   3648: 'Spare_Fault_3648', class No Acknowledgement, trigger "DB302_HMI_Faults_Carrier56_Faults_3" bit 15
   3649: 'Carrier 57 Disconnect Open Power Fault DI11.0', class No Acknowledgement, trigger "DB302_HMI_Faults_Carrier57_Faults_0" bit 0
   3650: 'Carrier 57 Drive Profinet Comm Fault', class No Acknowledgement, trigger "DB302_HMI_Faults_Carrier57_Faults_0" bit 1
   3651: 'Carrier 57 Production Stop Not Reset', class No Acknowledgement, trigger "DB302_HMI_Faults_Carrier57_Faults_0" bit 2
   3652: 'Carrier 57 CB02122 Tripped', class No Acknowledgement, trigger "DB302_HMI_Faults_Carrier57_Faults_0" bit 3
   3653: 'Carrier 57 CB02123 Tripped', class No Acknowledgement, trigger "DB302_HMI_Faults_Carrier57_Faults_0" bit 4
   3654: 'Carrier 57 AUX1 CB Tripped', class No Acknowledgement, trigger "DB302_HMI_Faults_Carrier57_Faults_0" bit 5
   3655: 'Carrier 57 AUX2 CB Tripped', class No Acknowledgement, trigger "DB302_HMI_Faults_Carrier57_Faults_0" bit 6
   3656: 'Carrier 57 PLC Not Communicating', class No Acknowledgement, trigger "DB302_HMI_Faults_Carrier57_Faults_0" bit 7
   3657: 'Carrier 57 Safe Input Card Fault', class No Acknowledgement, trigger "DB302_HMI_Faults_Carrier57_Faults_0" bit 8
   3658: 'Carrier 57 Safe Output Card Fault', class No Acknowledgement, trigger "DB302_HMI_Faults_Carrier57_Faults_0" bit 9
   3659: 'Carrier 57 Standard Input Card Fault', class No Acknowledgement, trigger "DB302_HMI_Faults_Carrier57_Faults_0" bit 10
   3660: 'Carrier 57 Standard Output Card Fault', class No Acknowledgement, trigger "DB302_HMI_Faults_Carrier57_Faults_0" bit 11
   3661: 'Carrier 57 Encoder Position Fault', class No Acknowledgement, trigger "DB302_HMI_Faults_Carrier57_Faults_0" bit 12
   3662: 'Carrier 57 Encoder Internal Error', class No Acknowledgement, trigger "DB302_HMI_Faults_Carrier57_Faults_0" bit 13
   3663: 'Carrier 57 Encoder Comm Fault', class No Acknowledgement, trigger "DB302_HMI_Faults_Carrier57_Faults_0" bit 14
   3664: 'Carrier 57 HMI Comm Fault', class No Acknowledgement, trigger "DB302_HMI_Faults_Carrier57_Faults_0" bit 15
   3665: 'Carrier 57 Crash Detection Fault', class No Acknowledgement, trigger "DB302_HMI_Faults_Carrier57_Faults_1" bit 0
   3666: 'Carrier 57 Carrier Number Invalid', class No Acknowledgement, trigger "DB302_HMI_Faults_Carrier57_Faults_1" bit 1
   3667: 'Carrier 57 Drive: PROFINET configuration error', class No Acknowledgement, trigger "DB302_HMI_Faults_Carrier57_Faults_1" bit 2
   3668: 'Carrier 57 Drive: Error internal communications', class No Acknowledgement, trigger "DB302_HMI_Faults_Carrier57_Faults_1" bit 3
   3669: 'Carrier 57 Drive: Motor overtemperature', class No Acknowledgement, trigger "DB302_HMI_Faults_Carrier57_Faults_1" bit 4
   3670: 'Carrier 57 Drive: Motor overcurrent', class No Acknowledgement, trigger "DB302_HMI_Faults_Carrier57_Faults_1" bit 5
   3671: 'Carrier 57 Drive: Infeed or power unit not ready', class No Acknowledgement, trigger "DB302_HMI_Faults_Carrier57_Faults_1" bit 6
   3672: 'Carrier 57 Drive: Short-circuit/ground fault detected', class No Acknowledgement, trigger "DB302_HMI_Faults_Carrier57_Faults_1" bit 7
   3673: 'Carrier 57 Drive: PROFINET Setpoint timeout', class No Acknowledgement, trigger "DB302_HMI_Faults_Carrier57_Faults_1" bit 8
   3674: 'Carrier 57 Power unit: Overcurrent', class No Acknowledgement, trigger "DB302_HMI_Faults_Carrier57_Faults_1" bit 9
   3675: 'Carrier 57 Power unit: DC link voltage overvoltage', class No Acknowledgement, trigger "DB302_HMI_Faults_Carrier57_Faults_1" bit 10
   3676: 'Carrier 57 Power unit: DC link voltage undervoltage', class No Acknowledgement, trigger "DB302_HMI_Faults_Carrier57_Faults_1" bit 11
   3677: 'Carrier 57 Power unit: Line phase failure in main circuit', class No Acknowledgement, trigger "DB302_HMI_Faults_Carrier57_Faults_1" bit 12
   3678: 'Carrier 57 Power unit: Phase failure motor cable', class No Acknowledgement, trigger "DB302_HMI_Faults_Carrier57_Faults_1" bit 13
   3679: 'Carrier 57 Power unit: Ground fault', class No Acknowledgement, trigger "DB302_HMI_Faults_Carrier57_Faults_1" bit 14
   3680: 'Spare_Fault_3680', class No Acknowledgement, trigger "DB302_HMI_Faults_Carrier57_Faults_1" bit 15
   3681: 'Carrier 57 Motion Off Fault', class No Acknowledgement, trigger "DB302_HMI_Faults_Carrier57_Faults_2" bit 0
   3682: 'Carrier 57 Motion On Fault', class No Acknowledgement, trigger "DB302_HMI_Faults_Carrier57_Faults_2" bit 1
   3683: 'Carrier 57 Spacing Fault', class No Acknowledgement, trigger "DB302_HMI_Faults_Carrier57_Faults_2" bit 2
   3684: 'Carrier 57 Duplicate Carrier Number Fault', class No Acknowledgement, trigger "DB302_HMI_Faults_Carrier57_Faults_2" bit 3
   3685: 'Spare_Fault_3685', class No Acknowledgement, trigger "DB302_HMI_Faults_Carrier57_Faults_2" bit 4
   3686: 'Spare_Fault_3686', class No Acknowledgement, trigger "DB302_HMI_Faults_Carrier57_Faults_2" bit 5
   3687: 'Spare_Fault_3687', class No Acknowledgement, trigger "DB302_HMI_Faults_Carrier57_Faults_2" bit 6
   3688: 'Spare_Fault_3688', class No Acknowledgement, trigger "DB302_HMI_Faults_Carrier57_Faults_2" bit 7
   3689: 'Spare_Fault_3689', class No Acknowledgement, trigger "DB302_HMI_Faults_Carrier57_Faults_2" bit 8
   3690: 'Spare_Fault_3690', class No Acknowledgement, trigger "DB302_HMI_Faults_Carrier57_Faults_2" bit 9
   3691: 'Spare_Fault_3691', class No Acknowledgement, trigger "DB302_HMI_Faults_Carrier57_Faults_2" bit 10
   3692: 'Spare_Fault_3692', class No Acknowledgement, trigger "DB302_HMI_Faults_Carrier57_Faults_2" bit 11
   3693: 'Spare_Fault_3693', class No Acknowledgement, trigger "DB302_HMI_Faults_Carrier57_Faults_2" bit 12
   3694: 'Spare_Fault_3694', class No Acknowledgement, trigger "DB302_HMI_Faults_Carrier57_Faults_2" bit 13
   3695: 'Spare_Fault_3695', class No Acknowledgement, trigger "DB302_HMI_Faults_Carrier57_Faults_2" bit 14
   3696: 'Spare_Fault_3696', class No Acknowledgement, trigger "DB302_HMI_Faults_Carrier57_Faults_2" bit 15
   3697: 'Spare_Fault_3697', class No Acknowledgement, trigger "DB302_HMI_Faults_Carrier57_Faults_3" bit 0
   3698: 'Spare_Fault_3698', class No Acknowledgement, trigger "DB302_HMI_Faults_Carrier57_Faults_3" bit 1
   3699: 'Spare_Fault_3699', class No Acknowledgement, trigger "DB302_HMI_Faults_Carrier57_Faults_3" bit 2
   3700: 'Spare_Fault_3700', class No Acknowledgement, trigger "DB302_HMI_Faults_Carrier57_Faults_3" bit 3
   3701: 'Spare_Fault_3701', class No Acknowledgement, trigger "DB302_HMI_Faults_Carrier57_Faults_3" bit 4
   3702: 'Spare_Fault_3702', class No Acknowledgement, trigger "DB302_HMI_Faults_Carrier57_Faults_3" bit 5
   3703: 'Spare_Fault_3703', class No Acknowledgement, trigger "DB302_HMI_Faults_Carrier57_Faults_3" bit 6
   3704: 'Spare_Fault_3704', class No Acknowledgement, trigger "DB302_HMI_Faults_Carrier57_Faults_3" bit 7
   3705: 'Spare_Fault_3705', class No Acknowledgement, trigger "DB302_HMI_Faults_Carrier57_Faults_3" bit 8
   3706: 'Spare_Fault_3706', class No Acknowledgement, trigger "DB302_HMI_Faults_Carrier57_Faults_3" bit 9
   3707: 'Spare_Fault_3707', class No Acknowledgement, trigger "DB302_HMI_Faults_Carrier57_Faults_3" bit 10
   3708: 'Spare_Fault_3708', class No Acknowledgement, trigger "DB302_HMI_Faults_Carrier57_Faults_3" bit 11
   3709: 'Spare_Fault_3709', class No Acknowledgement, trigger "DB302_HMI_Faults_Carrier57_Faults_3" bit 12
   3710: 'Spare_Fault_3710', class No Acknowledgement, trigger "DB302_HMI_Faults_Carrier57_Faults_3" bit 13
   3711: 'Spare_Fault_3711', class No Acknowledgement, trigger "DB302_HMI_Faults_Carrier57_Faults_3" bit 14
   3712: 'Spare_Fault_3712', class No Acknowledgement, trigger "DB302_HMI_Faults_Carrier57_Faults_3" bit 15
   3713: 'Carrier 58 Disconnect Open Power Fault DI11.0', class No Acknowledgement, trigger "DB302_HMI_Faults_Carrier58_Faults_0" bit 0
   3714: 'Carrier 58 Drive Profinet Comm Fault', class No Acknowledgement, trigger "DB302_HMI_Faults_Carrier58_Faults_0" bit 1
   3715: 'Carrier 58 Production Stop Not Reset', class No Acknowledgement, trigger "DB302_HMI_Faults_Carrier58_Faults_0" bit 2
   3716: 'Carrier 58 CB02122 Tripped', class No Acknowledgement, trigger "DB302_HMI_Faults_Carrier58_Faults_0" bit 3
   3717: 'Carrier 58 CB02123 Tripped', class No Acknowledgement, trigger "DB302_HMI_Faults_Carrier58_Faults_0" bit 4
   3718: 'Carrier 58 AUX1 CB Tripped', class No Acknowledgement, trigger "DB302_HMI_Faults_Carrier58_Faults_0" bit 5
   3719: 'Carrier 58 AUX2 CB Tripped', class No Acknowledgement, trigger "DB302_HMI_Faults_Carrier58_Faults_0" bit 6
   3720: 'Carrier 58 PLC Not Communicating', class No Acknowledgement, trigger "DB302_HMI_Faults_Carrier58_Faults_0" bit 7
   3721: 'Carrier 58 Safe Input Card Fault', class No Acknowledgement, trigger "DB302_HMI_Faults_Carrier58_Faults_0" bit 8
   3722: 'Carrier 58 Safe Output Card Fault', class No Acknowledgement, trigger "DB302_HMI_Faults_Carrier58_Faults_0" bit 9
   3723: 'Carrier 58 Standard Input Card Fault', class No Acknowledgement, trigger "DB302_HMI_Faults_Carrier58_Faults_0" bit 10
   3724: 'Carrier 58 Standard Output Card Fault', class No Acknowledgement, trigger "DB302_HMI_Faults_Carrier58_Faults_0" bit 11
   3725: 'Carrier 58 Encoder Position Fault', class No Acknowledgement, trigger "DB302_HMI_Faults_Carrier58_Faults_0" bit 12
   3726: 'Carrier 58 Encoder Internal Error', class No Acknowledgement, trigger "DB302_HMI_Faults_Carrier58_Faults_0" bit 13
   3727: 'Carrier 58 Encoder Comm Fault', class No Acknowledgement, trigger "DB302_HMI_Faults_Carrier58_Faults_0" bit 14
   3728: 'Carrier 58 HMI Comm Fault', class No Acknowledgement, trigger "DB302_HMI_Faults_Carrier58_Faults_0" bit 15
   3729: 'Carrier 58 Crash Detection Fault', class No Acknowledgement, trigger "DB302_HMI_Faults_Carrier58_Faults_1" bit 0
   3730: 'Carrier 58 Carrier Number Invalid', class No Acknowledgement, trigger "DB302_HMI_Faults_Carrier58_Faults_1" bit 1
   3731: 'Carrier 58 Drive: PROFINET configuration error', class No Acknowledgement, trigger "DB302_HMI_Faults_Carrier58_Faults_1" bit 2
   3732: 'Carrier 58 Drive: Error internal communications', class No Acknowledgement, trigger "DB302_HMI_Faults_Carrier58_Faults_1" bit 3
   3733: 'Carrier 58 Drive: Motor overtemperature', class No Acknowledgement, trigger "DB302_HMI_Faults_Carrier58_Faults_1" bit 4
   3734: 'Carrier 58 Drive: Motor overcurrent', class No Acknowledgement, trigger "DB302_HMI_Faults_Carrier58_Faults_1" bit 5
   3735: 'Carrier 58 Drive: Infeed or power unit not ready', class No Acknowledgement, trigger "DB302_HMI_Faults_Carrier58_Faults_1" bit 6
   3736: 'Carrier 58 Drive: Short-circuit/ground fault detected', class No Acknowledgement, trigger "DB302_HMI_Faults_Carrier58_Faults_1" bit 7
   3737: 'Carrier 58 Drive: PROFINET Setpoint timeout', class No Acknowledgement, trigger "DB302_HMI_Faults_Carrier58_Faults_1" bit 8
   3738: 'Carrier 58 Power unit: Overcurrent', class No Acknowledgement, trigger "DB302_HMI_Faults_Carrier58_Faults_1" bit 9
   3739: 'Carrier 58 Power unit: DC link voltage overvoltage', class No Acknowledgement, trigger "DB302_HMI_Faults_Carrier58_Faults_1" bit 10
   3740: 'Carrier 58 Power unit: DC link voltage undervoltage', class No Acknowledgement, trigger "DB302_HMI_Faults_Carrier58_Faults_1" bit 11
   3741: 'Carrier 58 Power unit: Line phase failure in main circuit', class No Acknowledgement, trigger "DB302_HMI_Faults_Carrier58_Faults_1" bit 12
   3742: 'Carrier 58 Power unit: Phase failure motor cable', class No Acknowledgement, trigger "DB302_HMI_Faults_Carrier58_Faults_1" bit 13
   3743: 'Carrier 58 Power unit: Ground fault', class No Acknowledgement, trigger "DB302_HMI_Faults_Carrier58_Faults_1" bit 14
   3744: 'Spare_Fault_3744', class No Acknowledgement, trigger "DB302_HMI_Faults_Carrier58_Faults_1" bit 15
   3745: 'Carrier 58 Motion Off Fault', class No Acknowledgement, trigger "DB302_HMI_Faults_Carrier58_Faults_2" bit 0
   3746: 'Carrier 58 Motion On Fault', class No Acknowledgement, trigger "DB302_HMI_Faults_Carrier58_Faults_2" bit 1
   3747: 'Carrier 58 Spacing Fault', class No Acknowledgement, trigger "DB302_HMI_Faults_Carrier58_Faults_2" bit 2
   3748: 'Carrier 58 Duplicate Carrier Number Fault', class No Acknowledgement, trigger "DB302_HMI_Faults_Carrier58_Faults_2" bit 3
   3749: 'Spare_Fault_3749', class No Acknowledgement, trigger "DB302_HMI_Faults_Carrier58_Faults_2" bit 4
   3750: 'Spare_Fault_3750', class No Acknowledgement, trigger "DB302_HMI_Faults_Carrier58_Faults_2" bit 5
   3751: 'Spare_Fault_3751', class No Acknowledgement, trigger "DB302_HMI_Faults_Carrier58_Faults_2" bit 6
   3752: 'Spare_Fault_3752', class No Acknowledgement, trigger "DB302_HMI_Faults_Carrier58_Faults_2" bit 7
   3753: 'Spare_Fault_3753', class No Acknowledgement, trigger "DB302_HMI_Faults_Carrier58_Faults_2" bit 8
   3754: 'Spare_Fault_3754', class No Acknowledgement, trigger "DB302_HMI_Faults_Carrier58_Faults_2" bit 9
   3755: 'Spare_Fault_3755', class No Acknowledgement, trigger "DB302_HMI_Faults_Carrier58_Faults_2" bit 10
   3756: 'Spare_Fault_3756', class No Acknowledgement, trigger "DB302_HMI_Faults_Carrier58_Faults_2" bit 11
   3757: 'Spare_Fault_3757', class No Acknowledgement, trigger "DB302_HMI_Faults_Carrier58_Faults_2" bit 12
   3758: 'Spare_Fault_3758', class No Acknowledgement, trigger "DB302_HMI_Faults_Carrier58_Faults_2" bit 13
   3759: 'Spare_Fault_3759', class No Acknowledgement, trigger "DB302_HMI_Faults_Carrier58_Faults_2" bit 14
   3760: 'Spare_Fault_3760', class No Acknowledgement, trigger "DB302_HMI_Faults_Carrier58_Faults_2" bit 15
   3761: 'Spare_Fault_3761', class No Acknowledgement, trigger "DB302_HMI_Faults_Carrier58_Faults_3" bit 0
   3762: 'Spare_Fault_3762', class No Acknowledgement, trigger "DB302_HMI_Faults_Carrier58_Faults_3" bit 1
   3763: 'Spare_Fault_3763', class No Acknowledgement, trigger "DB302_HMI_Faults_Carrier58_Faults_3" bit 2
   3764: 'Spare_Fault_3764', class No Acknowledgement, trigger "DB302_HMI_Faults_Carrier58_Faults_3" bit 3
   3765: 'Spare_Fault_3765', class No Acknowledgement, trigger "DB302_HMI_Faults_Carrier58_Faults_3" bit 4
   3766: 'Spare_Fault_3766', class No Acknowledgement, trigger "DB302_HMI_Faults_Carrier58_Faults_3" bit 5
   3767: 'Spare_Fault_3767', class No Acknowledgement, trigger "DB302_HMI_Faults_Carrier58_Faults_3" bit 6
   3768: 'Spare_Fault_3768', class No Acknowledgement, trigger "DB302_HMI_Faults_Carrier58_Faults_3" bit 7
   3769: 'Spare_Fault_3769', class No Acknowledgement, trigger "DB302_HMI_Faults_Carrier58_Faults_3" bit 8
   3770: 'Spare_Fault_3770', class No Acknowledgement, trigger "DB302_HMI_Faults_Carrier58_Faults_3" bit 9
   3771: 'Spare_Fault_3771', class No Acknowledgement, trigger "DB302_HMI_Faults_Carrier58_Faults_3" bit 10
   3772: 'Spare_Fault_3772', class No Acknowledgement, trigger "DB302_HMI_Faults_Carrier58_Faults_3" bit 11
   3773: 'Spare_Fault_3773', class No Acknowledgement, trigger "DB302_HMI_Faults_Carrier58_Faults_3" bit 12
   3774: 'Spare_Fault_3774', class No Acknowledgement, trigger "DB302_HMI_Faults_Carrier58_Faults_3" bit 13
   3775: 'Spare_Fault_3775', class No Acknowledgement, trigger "DB302_HMI_Faults_Carrier58_Faults_3" bit 14
   3776: 'Spare_Fault_3776', class No Acknowledgement, trigger "DB302_HMI_Faults_Carrier58_Faults_3" bit 15
   3777: 'Carrier 59 Disconnect Open Power Fault DI11.0', class No Acknowledgement, trigger "DB302_HMI_Faults_Carrier59_Faults_0" bit 0
   3778: 'Carrier 59 Drive Profinet Comm Fault', class No Acknowledgement, trigger "DB302_HMI_Faults_Carrier59_Faults_0" bit 1
   3779: 'Carrier 59 Production Stop Not Reset', class No Acknowledgement, trigger "DB302_HMI_Faults_Carrier59_Faults_0" bit 2
   3780: 'Carrier 59 CB02122 Tripped', class No Acknowledgement, trigger "DB302_HMI_Faults_Carrier59_Faults_0" bit 3
   3781: 'Carrier 59 CB02123 Tripped', class No Acknowledgement, trigger "DB302_HMI_Faults_Carrier59_Faults_0" bit 4
   3782: 'Carrier 59 AUX1 CB Tripped', class No Acknowledgement, trigger "DB302_HMI_Faults_Carrier59_Faults_0" bit 5
   3783: 'Carrier 59 AUX2 CB Tripped', class No Acknowledgement, trigger "DB302_HMI_Faults_Carrier59_Faults_0" bit 6
   3784: 'Carrier 59 PLC Not Communicating', class No Acknowledgement, trigger "DB302_HMI_Faults_Carrier59_Faults_0" bit 7
   3785: 'Carrier 59 Safe Input Card Fault', class No Acknowledgement, trigger "DB302_HMI_Faults_Carrier59_Faults_0" bit 8
   3786: 'Carrier 59 Safe Output Card Fault', class No Acknowledgement, trigger "DB302_HMI_Faults_Carrier59_Faults_0" bit 9
   3787: 'Carrier 59 Standard Input Card Fault', class No Acknowledgement, trigger "DB302_HMI_Faults_Carrier59_Faults_0" bit 10
   3788: 'Carrier 59 Standard Output Card Fault', class No Acknowledgement, trigger "DB302_HMI_Faults_Carrier59_Faults_0" bit 11
   3789: 'Carrier 59 Encoder Position Fault', class No Acknowledgement, trigger "DB302_HMI_Faults_Carrier59_Faults_0" bit 12
   3790: 'Carrier 59 Encoder Internal Error', class No Acknowledgement, trigger "DB302_HMI_Faults_Carrier59_Faults_0" bit 13
   3791: 'Carrier 59 Encoder Comm Fault', class No Acknowledgement, trigger "DB302_HMI_Faults_Carrier59_Faults_0" bit 14
   3792: 'Carrier 59 HMI Comm Fault', class No Acknowledgement, trigger "DB302_HMI_Faults_Carrier59_Faults_0" bit 15
   3793: 'Carrier 59 Crash Detection Fault', class No Acknowledgement, trigger "DB302_HMI_Faults_Carrier59_Faults_1" bit 0
   3794: 'Carrier 59 Carrier Number Invalid', class No Acknowledgement, trigger "DB302_HMI_Faults_Carrier59_Faults_1" bit 1
   3795: 'Carrier 59 Drive: PROFINET configuration error', class No Acknowledgement, trigger "DB302_HMI_Faults_Carrier59_Faults_1" bit 2
   3796: 'Carrier 59 Drive: Error internal communications', class No Acknowledgement, trigger "DB302_HMI_Faults_Carrier59_Faults_1" bit 3
   3797: 'Carrier 59 Drive: Motor overtemperature', class No Acknowledgement, trigger "DB302_HMI_Faults_Carrier59_Faults_1" bit 4
   3798: 'Carrier 59 Drive: Motor overcurrent', class No Acknowledgement, trigger "DB302_HMI_Faults_Carrier59_Faults_1" bit 5
   3799: 'Carrier 59 Drive: Infeed or power unit not ready', class No Acknowledgement, trigger "DB302_HMI_Faults_Carrier59_Faults_1" bit 6
   3800: 'Carrier 59 Drive: Short-circuit/ground fault detected', class No Acknowledgement, trigger "DB302_HMI_Faults_Carrier59_Faults_1" bit 7
   3801: 'Carrier 59 Drive: PROFINET Setpoint timeout', class No Acknowledgement, trigger "DB302_HMI_Faults_Carrier59_Faults_1" bit 8
   3802: 'Carrier 59 Power unit: Overcurrent', class No Acknowledgement, trigger "DB302_HMI_Faults_Carrier59_Faults_1" bit 9
   3803: 'Carrier 59 Power unit: DC link voltage overvoltage', class No Acknowledgement, trigger "DB302_HMI_Faults_Carrier59_Faults_1" bit 10
   3804: 'Carrier 59 Power unit: DC link voltage undervoltage', class No Acknowledgement, trigger "DB302_HMI_Faults_Carrier59_Faults_1" bit 11
   3805: 'Carrier 59 Power unit: Line phase failure in main circuit', class No Acknowledgement, trigger "DB302_HMI_Faults_Carrier59_Faults_1" bit 12
   3806: 'Carrier 59 Power unit: Phase failure motor cable', class No Acknowledgement, trigger "DB302_HMI_Faults_Carrier59_Faults_1" bit 13
   3807: 'Carrier 59 Power unit: Ground fault', class No Acknowledgement, trigger "DB302_HMI_Faults_Carrier59_Faults_1" bit 14
   3808: 'Spare_Fault_3808', class No Acknowledgement, trigger "DB302_HMI_Faults_Carrier59_Faults_1" bit 15
   3809: 'Carrier 59 Motion Off Fault', class No Acknowledgement, trigger "DB302_HMI_Faults_Carrier59_Faults_2" bit 0
   3810: 'Carrier 59 Motion On Fault', class No Acknowledgement, trigger "DB302_HMI_Faults_Carrier59_Faults_2" bit 1
   3811: 'Carrier 59 Spacing Fault', class No Acknowledgement, trigger "DB302_HMI_Faults_Carrier59_Faults_2" bit 2
   3812: 'Carrier 59 Duplicate Carrier Number Fault', class No Acknowledgement, trigger "DB302_HMI_Faults_Carrier59_Faults_2" bit 3
   3813: 'Spare_Fault_3813', class No Acknowledgement, trigger "DB302_HMI_Faults_Carrier59_Faults_2" bit 4
   3814: 'Spare_Fault_3814', class No Acknowledgement, trigger "DB302_HMI_Faults_Carrier59_Faults_2" bit 5
   3815: 'Spare_Fault_3815', class No Acknowledgement, trigger "DB302_HMI_Faults_Carrier59_Faults_2" bit 6
   3816: 'Spare_Fault_3816', class No Acknowledgement, trigger "DB302_HMI_Faults_Carrier59_Faults_2" bit 7
   3817: 'Spare_Fault_3817', class No Acknowledgement, trigger "DB302_HMI_Faults_Carrier59_Faults_2" bit 8
   3818: 'Spare_Fault_3818', class No Acknowledgement, trigger "DB302_HMI_Faults_Carrier59_Faults_2" bit 9
   3819: 'Spare_Fault_3819', class No Acknowledgement, trigger "DB302_HMI_Faults_Carrier59_Faults_2" bit 10
   3820: 'Spare_Fault_3820', class No Acknowledgement, trigger "DB302_HMI_Faults_Carrier59_Faults_2" bit 11
   3821: 'Spare_Fault_3821', class No Acknowledgement, trigger "DB302_HMI_Faults_Carrier59_Faults_2" bit 12
   3822: 'Spare_Fault_3822', class No Acknowledgement, trigger "DB302_HMI_Faults_Carrier59_Faults_2" bit 13
   3823: 'Spare_Fault_3823', class No Acknowledgement, trigger "DB302_HMI_Faults_Carrier59_Faults_2" bit 14
   3824: 'Spare_Fault_3824', class No Acknowledgement, trigger "DB302_HMI_Faults_Carrier59_Faults_2" bit 15
   3825: 'Spare_Fault_3825', class No Acknowledgement, trigger "DB302_HMI_Faults_Carrier59_Faults_3" bit 0
   3826: 'Spare_Fault_3826', class No Acknowledgement, trigger "DB302_HMI_Faults_Carrier59_Faults_3" bit 1
   3827: 'Spare_Fault_3827', class No Acknowledgement, trigger "DB302_HMI_Faults_Carrier59_Faults_3" bit 2
   3828: 'Spare_Fault_3828', class No Acknowledgement, trigger "DB302_HMI_Faults_Carrier59_Faults_3" bit 3
   3829: 'Spare_Fault_3829', class No Acknowledgement, trigger "DB302_HMI_Faults_Carrier59_Faults_3" bit 4
   3830: 'Spare_Fault_3830', class No Acknowledgement, trigger "DB302_HMI_Faults_Carrier59_Faults_3" bit 5
   3831: 'Spare_Fault_3831', class No Acknowledgement, trigger "DB302_HMI_Faults_Carrier59_Faults_3" bit 6
   3832: 'Spare_Fault_3832', class No Acknowledgement, trigger "DB302_HMI_Faults_Carrier59_Faults_3" bit 7
   3833: 'Spare_Fault_3833', class No Acknowledgement, trigger "DB302_HMI_Faults_Carrier59_Faults_3" bit 8
   3834: 'Spare_Fault_3834', class No Acknowledgement, trigger "DB302_HMI_Faults_Carrier59_Faults_3" bit 9
   3835: 'Spare_Fault_3835', class No Acknowledgement, trigger "DB302_HMI_Faults_Carrier59_Faults_3" bit 10
   3836: 'Spare_Fault_3836', class No Acknowledgement, trigger "DB302_HMI_Faults_Carrier59_Faults_3" bit 11
   3837: 'Spare_Fault_3837', class No Acknowledgement, trigger "DB302_HMI_Faults_Carrier59_Faults_3" bit 12
   3838: 'Spare_Fault_3838', class No Acknowledgement, trigger "DB302_HMI_Faults_Carrier59_Faults_3" bit 13
   3839: 'Spare_Fault_3839', class No Acknowledgement, trigger "DB302_HMI_Faults_Carrier59_Faults_3" bit 14
   3840: 'Spare_Fault_3840', class No Acknowledgement, trigger "DB302_HMI_Faults_Carrier59_Faults_3" bit 15
   3841: 'Carrier 60 Disconnect Open Power Fault DI11.0', class No Acknowledgement, trigger "DB302_HMI_Faults_Carrier60_Faults_0" bit 0
   3842: 'Carrier 60 Drive Profinet Comm Fault', class No Acknowledgement, trigger "DB302_HMI_Faults_Carrier60_Faults_0" bit 1
   3843: 'Carrier 60 Production Stop Not Reset', class No Acknowledgement, trigger "DB302_HMI_Faults_Carrier60_Faults_0" bit 2
   3844: 'Carrier 60 CB02122 Tripped', class No Acknowledgement, trigger "DB302_HMI_Faults_Carrier60_Faults_0" bit 3
   3845: 'Carrier 60 CB02123 Tripped', class No Acknowledgement, trigger "DB302_HMI_Faults_Carrier60_Faults_0" bit 4
   3846: 'Carrier 60 AUX1 CB Tripped', class No Acknowledgement, trigger "DB302_HMI_Faults_Carrier60_Faults_0" bit 5
   3847: 'Carrier 60 AUX2 CB Tripped', class No Acknowledgement, trigger "DB302_HMI_Faults_Carrier60_Faults_0" bit 6
   3848: 'Carrier 60 PLC Not Communicating', class No Acknowledgement, trigger "DB302_HMI_Faults_Carrier60_Faults_0" bit 7
   3849: 'Carrier 60 Safe Input Card Fault', class No Acknowledgement, trigger "DB302_HMI_Faults_Carrier60_Faults_0" bit 8
   3850: 'Carrier 60 Safe Output Card Fault', class No Acknowledgement, trigger "DB302_HMI_Faults_Carrier60_Faults_0" bit 9
   3851: 'Carrier 60 Standard Input Card Fault', class No Acknowledgement, trigger "DB302_HMI_Faults_Carrier60_Faults_0" bit 10
   3852: 'Carrier 60 Standard Output Card Fault', class No Acknowledgement, trigger "DB302_HMI_Faults_Carrier60_Faults_0" bit 11
   3853: 'Carrier 60 Encoder Position Fault', class No Acknowledgement, trigger "DB302_HMI_Faults_Carrier60_Faults_0" bit 12
   3854: 'Carrier 60 Encoder Internal Error', class No Acknowledgement, trigger "DB302_HMI_Faults_Carrier60_Faults_0" bit 13
   3855: 'Carrier 60 Encoder Comm Fault', class No Acknowledgement, trigger "DB302_HMI_Faults_Carrier60_Faults_0" bit 14
   3856: 'Carrier 60 HMI Comm Fault', class No Acknowledgement, trigger "DB302_HMI_Faults_Carrier60_Faults_0" bit 15
   3857: 'Carrier 60 Crash Detection Fault', class No Acknowledgement, trigger "DB302_HMI_Faults_Carrier60_Faults_1" bit 0
   3858: 'Carrier 60 Carrier Number Invalid', class No Acknowledgement, trigger "DB302_HMI_Faults_Carrier60_Faults_1" bit 1
   3859: 'Carrier 60 Drive: PROFINET configuration error', class No Acknowledgement, trigger "DB302_HMI_Faults_Carrier60_Faults_1" bit 2
   3860: 'Carrier 60 Drive: Error internal communications', class No Acknowledgement, trigger "DB302_HMI_Faults_Carrier60_Faults_1" bit 3
   3861: 'Carrier 60 Drive: Motor overtemperature', class No Acknowledgement, trigger "DB302_HMI_Faults_Carrier60_Faults_1" bit 4
   3862: 'Carrier 60 Drive: Motor overcurrent', class No Acknowledgement, trigger "DB302_HMI_Faults_Carrier60_Faults_1" bit 5
   3863: 'Carrier 60 Drive: Infeed or power unit not ready', class No Acknowledgement, trigger "DB302_HMI_Faults_Carrier60_Faults_1" bit 6
   3864: 'Carrier 60 Drive: Short-circuit/ground fault detected', class No Acknowledgement, trigger "DB302_HMI_Faults_Carrier60_Faults_1" bit 7
   3865: 'Carrier 60 Drive: PROFINET Setpoint timeout', class No Acknowledgement, trigger "DB302_HMI_Faults_Carrier60_Faults_1" bit 8
   3866: 'Carrier 60 Power unit: Overcurrent', class No Acknowledgement, trigger "DB302_HMI_Faults_Carrier60_Faults_1" bit 9
   3867: 'Carrier 60 Power unit: DC link voltage overvoltage', class No Acknowledgement, trigger "DB302_HMI_Faults_Carrier60_Faults_1" bit 10
   3868: 'Carrier 60 Power unit: DC link voltage undervoltage', class No Acknowledgement, trigger "DB302_HMI_Faults_Carrier60_Faults_1" bit 11
   3869: 'Carrier 60 Power unit: Line phase failure in main circuit', class No Acknowledgement, trigger "DB302_HMI_Faults_Carrier60_Faults_1" bit 12
   3870: 'Carrier 60 Power unit: Phase failure motor cable', class No Acknowledgement, trigger "DB302_HMI_Faults_Carrier60_Faults_1" bit 13
   3871: 'Carrier 60 Power unit: Ground fault', class No Acknowledgement, trigger "DB302_HMI_Faults_Carrier60_Faults_1" bit 14
   3872: 'Spare_Fault_3872', class No Acknowledgement, trigger "DB302_HMI_Faults_Carrier60_Faults_1" bit 15
   3873: 'Carrier 60 Motion Off Fault', class No Acknowledgement, trigger "DB302_HMI_Faults_Carrier60_Faults_2" bit 0
   3874: 'Carrier 60 Motion On Fault', class No Acknowledgement, trigger "DB302_HMI_Faults_Carrier60_Faults_2" bit 1
   3875: 'Carrier 60 Spacing Fault', class No Acknowledgement, trigger "DB302_HMI_Faults_Carrier60_Faults_2" bit 2
   3876: 'Carrier 60 Duplicate Carrier Number Fault', class No Acknowledgement, trigger "DB302_HMI_Faults_Carrier60_Faults_2" bit 3
   3877: 'Spare_Fault_3877', class No Acknowledgement, trigger "DB302_HMI_Faults_Carrier60_Faults_2" bit 4
   3878: 'Spare_Fault_3878', class No Acknowledgement, trigger "DB302_HMI_Faults_Carrier60_Faults_2" bit 5
   3879: 'Spare_Fault_3879', class No Acknowledgement, trigger "DB302_HMI_Faults_Carrier60_Faults_2" bit 6
   3880: 'Spare_Fault_3880', class No Acknowledgement, trigger "DB302_HMI_Faults_Carrier60_Faults_2" bit 7
   3881: 'Spare_Fault_3881', class No Acknowledgement, trigger "DB302_HMI_Faults_Carrier60_Faults_2" bit 8
   3882: 'Spare_Fault_3882', class No Acknowledgement, trigger "DB302_HMI_Faults_Carrier60_Faults_2" bit 9
   3883: 'Spare_Fault_3883', class No Acknowledgement, trigger "DB302_HMI_Faults_Carrier60_Faults_2" bit 10
   3884: 'Spare_Fault_3884', class No Acknowledgement, trigger "DB302_HMI_Faults_Carrier60_Faults_2" bit 11
   3885: 'Spare_Fault_3885', class No Acknowledgement, trigger "DB302_HMI_Faults_Carrier60_Faults_2" bit 12
   3886: 'Spare_Fault_3886', class No Acknowledgement, trigger "DB302_HMI_Faults_Carrier60_Faults_2" bit 13
   3887: 'Spare_Fault_3887', class No Acknowledgement, trigger "DB302_HMI_Faults_Carrier60_Faults_2" bit 14
   3888: 'Spare_Fault_3888', class No Acknowledgement, trigger "DB302_HMI_Faults_Carrier60_Faults_2" bit 15
   3889: 'Spare_Fault_3889', class No Acknowledgement, trigger "DB302_HMI_Faults_Carrier60_Faults_3" bit 0
   3890: 'Spare_Fault_3890', class No Acknowledgement, trigger "DB302_HMI_Faults_Carrier60_Faults_3" bit 1
   3891: 'Spare_Fault_3891', class No Acknowledgement, trigger "DB302_HMI_Faults_Carrier60_Faults_3" bit 2
   3892: 'Spare_Fault_3892', class No Acknowledgement, trigger "DB302_HMI_Faults_Carrier60_Faults_3" bit 3
   3893: 'Spare_Fault_3893', class No Acknowledgement, trigger "DB302_HMI_Faults_Carrier60_Faults_3" bit 4
   3894: 'Spare_Fault_3894', class No Acknowledgement, trigger "DB302_HMI_Faults_Carrier60_Faults_3" bit 5
   3895: 'Spare_Fault_3895', class No Acknowledgement, trigger "DB302_HMI_Faults_Carrier60_Faults_3" bit 6
   3896: 'Spare_Fault_3896', class No Acknowledgement, trigger "DB302_HMI_Faults_Carrier60_Faults_3" bit 7
   3897: 'Spare_Fault_3897', class No Acknowledgement, trigger "DB302_HMI_Faults_Carrier60_Faults_3" bit 8
   3898: 'Spare_Fault_3898', class No Acknowledgement, trigger "DB302_HMI_Faults_Carrier60_Faults_3" bit 9
   3899: 'Spare_Fault_3899', class No Acknowledgement, trigger "DB302_HMI_Faults_Carrier60_Faults_3" bit 10
   3900: 'Spare_Fault_3900', class No Acknowledgement, trigger "DB302_HMI_Faults_Carrier60_Faults_3" bit 11
   3901: 'Spare_Fault_3901', class No Acknowledgement, trigger "DB302_HMI_Faults_Carrier60_Faults_3" bit 12
   3902: 'Spare_Fault_3902', class No Acknowledgement, trigger "DB302_HMI_Faults_Carrier60_Faults_3" bit 13
   3903: 'Spare_Fault_3903', class No Acknowledgement, trigger "DB302_HMI_Faults_Carrier60_Faults_3" bit 14
   3904: 'Spare_Fault_3904', class No Acknowledgement, trigger "DB302_HMI_Faults_Carrier60_Faults_3" bit 15
   3905: 'Carrier 61 Disconnect Open Power Fault DI11.0', class No Acknowledgement, trigger "DB302_HMI_Faults_Carrier61_Faults_0" bit 0
   3906: 'Carrier 61 Drive Profinet Comm Fault', class No Acknowledgement, trigger "DB302_HMI_Faults_Carrier61_Faults_0" bit 1
   3907: 'Carrier 61 Production Stop Not Reset', class No Acknowledgement, trigger "DB302_HMI_Faults_Carrier61_Faults_0" bit 2
   3908: 'Carrier 61 CB02122 Tripped', class No Acknowledgement, trigger "DB302_HMI_Faults_Carrier61_Faults_0" bit 3
   3909: 'Carrier 61 CB02123 Tripped', class No Acknowledgement, trigger "DB302_HMI_Faults_Carrier61_Faults_0" bit 4
   3910: 'Carrier 61 AUX1 CB Tripped', class No Acknowledgement, trigger "DB302_HMI_Faults_Carrier61_Faults_0" bit 5
   3911: 'Carrier 61 AUX2 CB Tripped', class No Acknowledgement, trigger "DB302_HMI_Faults_Carrier61_Faults_0" bit 6
   3912: 'Carrier 61 PLC Not Communicating', class No Acknowledgement, trigger "DB302_HMI_Faults_Carrier61_Faults_0" bit 7
   3913: 'Carrier 61 Safe Input Card Fault', class No Acknowledgement, trigger "DB302_HMI_Faults_Carrier61_Faults_0" bit 8
   3914: 'Carrier 61 Safe Output Card Fault', class No Acknowledgement, trigger "DB302_HMI_Faults_Carrier61_Faults_0" bit 9
   3915: 'Carrier 61 Standard Input Card Fault', class No Acknowledgement, trigger "DB302_HMI_Faults_Carrier61_Faults_0" bit 10
   3916: 'Carrier 61 Standard Output Card Fault', class No Acknowledgement, trigger "DB302_HMI_Faults_Carrier61_Faults_0" bit 11
   3917: 'Carrier 61 Encoder Position Fault', class No Acknowledgement, trigger "DB302_HMI_Faults_Carrier61_Faults_0" bit 12
   3918: 'Carrier 61 Encoder Internal Error', class No Acknowledgement, trigger "DB302_HMI_Faults_Carrier61_Faults_0" bit 13
   3919: 'Carrier 61 Encoder Comm Fault', class No Acknowledgement, trigger "DB302_HMI_Faults_Carrier61_Faults_0" bit 14
   3920: 'Carrier 61 HMI Comm Fault', class No Acknowledgement, trigger "DB302_HMI_Faults_Carrier61_Faults_0" bit 15
   3921: 'Carrier 61 Crash Detection Fault', class No Acknowledgement, trigger "DB302_HMI_Faults_Carrier61_Faults_1" bit 0
   3922: 'Carrier 61 Carrier Number Invalid', class No Acknowledgement, trigger "DB302_HMI_Faults_Carrier61_Faults_1" bit 1
   3923: 'Carrier 61 Drive: PROFINET configuration error', class No Acknowledgement, trigger "DB302_HMI_Faults_Carrier61_Faults_1" bit 2
   3924: 'Carrier 61 Drive: Error internal communications', class No Acknowledgement, trigger "DB302_HMI_Faults_Carrier61_Faults_1" bit 3
   3925: 'Carrier 61 Drive: Motor overtemperature', class No Acknowledgement, trigger "DB302_HMI_Faults_Carrier61_Faults_1" bit 4
   3926: 'Carrier 61 Drive: Motor overcurrent', class No Acknowledgement, trigger "DB302_HMI_Faults_Carrier61_Faults_1" bit 5
   3927: 'Carrier 61 Drive: Infeed or power unit not ready', class No Acknowledgement, trigger "DB302_HMI_Faults_Carrier61_Faults_1" bit 6
   3928: 'Carrier 61 Drive: Short-circuit/ground fault detected', class No Acknowledgement, trigger "DB302_HMI_Faults_Carrier61_Faults_1" bit 7
   3929: 'Carrier 61 Drive: PROFINET Setpoint timeout', class No Acknowledgement, trigger "DB302_HMI_Faults_Carrier61_Faults_1" bit 8
   3930: 'Carrier 61 Power unit: Overcurrent', class No Acknowledgement, trigger "DB302_HMI_Faults_Carrier61_Faults_1" bit 9
   3931: 'Carrier 61 Power unit: DC link voltage overvoltage', class No Acknowledgement, trigger "DB302_HMI_Faults_Carrier61_Faults_1" bit 10
   3932: 'Carrier 61 Power unit: DC link voltage undervoltage', class No Acknowledgement, trigger "DB302_HMI_Faults_Carrier61_Faults_1" bit 11
   3933: 'Carrier 61 Power unit: Line phase failure in main circuit', class No Acknowledgement, trigger "DB302_HMI_Faults_Carrier61_Faults_1" bit 12
   3934: 'Carrier 61 Power unit: Phase failure motor cable', class No Acknowledgement, trigger "DB302_HMI_Faults_Carrier61_Faults_1" bit 13
   3935: 'Carrier 61 Power unit: Ground fault', class No Acknowledgement, trigger "DB302_HMI_Faults_Carrier61_Faults_1" bit 14
   3936: 'Spare_Fault_3936', class No Acknowledgement, trigger "DB302_HMI_Faults_Carrier61_Faults_1" bit 15
   3937: 'Carrier 61 Motion Off Fault', class No Acknowledgement, trigger "DB302_HMI_Faults_Carrier61_Faults_2" bit 0
   3938: 'Carrier 61 Motion On Fault', class No Acknowledgement, trigger "DB302_HMI_Faults_Carrier61_Faults_2" bit 1
   3939: 'Carrier 61 Spacing Fault', class No Acknowledgement, trigger "DB302_HMI_Faults_Carrier61_Faults_2" bit 2
   3940: 'Carrier 61 Duplicate Carrier Number Fault', class No Acknowledgement, trigger "DB302_HMI_Faults_Carrier61_Faults_2" bit 3
   3941: 'Spare_Fault_3941', class No Acknowledgement, trigger "DB302_HMI_Faults_Carrier61_Faults_2" bit 4
   3942: 'Spare_Fault_3942', class No Acknowledgement, trigger "DB302_HMI_Faults_Carrier61_Faults_2" bit 5
   3943: 'Spare_Fault_3943', class No Acknowledgement, trigger "DB302_HMI_Faults_Carrier61_Faults_2" bit 6
   3944: 'Spare_Fault_3944', class No Acknowledgement, trigger "DB302_HMI_Faults_Carrier61_Faults_2" bit 7
   3945: 'Spare_Fault_3945', class No Acknowledgement, trigger "DB302_HMI_Faults_Carrier61_Faults_2" bit 8
   3946: 'Spare_Fault_3946', class No Acknowledgement, trigger "DB302_HMI_Faults_Carrier61_Faults_2" bit 9
   3947: 'Spare_Fault_3947', class No Acknowledgement, trigger "DB302_HMI_Faults_Carrier61_Faults_2" bit 10
   3948: 'Spare_Fault_3948', class No Acknowledgement, trigger "DB302_HMI_Faults_Carrier61_Faults_2" bit 11
   3949: 'Spare_Fault_3949', class No Acknowledgement, trigger "DB302_HMI_Faults_Carrier61_Faults_2" bit 12
   3950: 'Spare_Fault_3950', class No Acknowledgement, trigger "DB302_HMI_Faults_Carrier61_Faults_2" bit 13
   3951: 'Spare_Fault_3951', class No Acknowledgement, trigger "DB302_HMI_Faults_Carrier61_Faults_2" bit 14
   3952: 'Spare_Fault_3952', class No Acknowledgement, trigger "DB302_HMI_Faults_Carrier61_Faults_2" bit 15
   3953: 'Spare_Fault_3953', class No Acknowledgement, trigger "DB302_HMI_Faults_Carrier61_Faults_3" bit 0
   3954: 'Spare_Fault_3954', class No Acknowledgement, trigger "DB302_HMI_Faults_Carrier61_Faults_3" bit 1
   3955: 'Spare_Fault_3955', class No Acknowledgement, trigger "DB302_HMI_Faults_Carrier61_Faults_3" bit 2
   3956: 'Spare_Fault_3956', class No Acknowledgement, trigger "DB302_HMI_Faults_Carrier61_Faults_3" bit 3
   3957: 'Spare_Fault_3957', class No Acknowledgement, trigger "DB302_HMI_Faults_Carrier61_Faults_3" bit 4
   3958: 'Spare_Fault_3958', class No Acknowledgement, trigger "DB302_HMI_Faults_Carrier61_Faults_3" bit 5
   3959: 'Spare_Fault_3959', class No Acknowledgement, trigger "DB302_HMI_Faults_Carrier61_Faults_3" bit 6
   3960: 'Spare_Fault_3960', class No Acknowledgement, trigger "DB302_HMI_Faults_Carrier61_Faults_3" bit 7
   3961: 'Spare_Fault_3961', class No Acknowledgement, trigger "DB302_HMI_Faults_Carrier61_Faults_3" bit 8
   3962: 'Spare_Fault_3962', class No Acknowledgement, trigger "DB302_HMI_Faults_Carrier61_Faults_3" bit 9
   3963: 'Spare_Fault_3963', class No Acknowledgement, trigger "DB302_HMI_Faults_Carrier61_Faults_3" bit 10
   3964: 'Spare_Fault_3964', class No Acknowledgement, trigger "DB302_HMI_Faults_Carrier61_Faults_3" bit 11
   3965: 'Spare_Fault_3965', class No Acknowledgement, trigger "DB302_HMI_Faults_Carrier61_Faults_3" bit 12
   3966: 'Spare_Fault_3966', class No Acknowledgement, trigger "DB302_HMI_Faults_Carrier61_Faults_3" bit 13
   3967: 'Spare_Fault_3967', class No Acknowledgement, trigger "DB302_HMI_Faults_Carrier61_Faults_3" bit 14
   3968: 'Spare_Fault_3968', class No Acknowledgement, trigger "DB302_HMI_Faults_Carrier61_Faults_3" bit 15
   3969: 'Carrier 62 Disconnect Open Power Fault DI11.0', class No Acknowledgement, trigger "DB302_HMI_Faults_Carrier62_Faults_0" bit 0
   3970: 'Carrier 62 Drive Profinet Comm Fault', class No Acknowledgement, trigger "DB302_HMI_Faults_Carrier62_Faults_0" bit 1
   3971: 'Carrier 62 Production Stop Not Reset', class No Acknowledgement, trigger "DB302_HMI_Faults_Carrier62_Faults_0" bit 2
   3972: 'Carrier 62 CB02122 Tripped', class No Acknowledgement, trigger "DB302_HMI_Faults_Carrier62_Faults_0" bit 3
   3973: 'Carrier 62 CB02123 Tripped', class No Acknowledgement, trigger "DB302_HMI_Faults_Carrier62_Faults_0" bit 4
   3974: 'Carrier 62 AUX1 CB Tripped', class No Acknowledgement, trigger "DB302_HMI_Faults_Carrier62_Faults_0" bit 5
   3975: 'Carrier 62 AUX2 CB Tripped', class No Acknowledgement, trigger "DB302_HMI_Faults_Carrier62_Faults_0" bit 6
   3976: 'Carrier 62 PLC Not Communicating', class No Acknowledgement, trigger "DB302_HMI_Faults_Carrier62_Faults_0" bit 7
   3977: 'Carrier 62 Safe Input Card Fault', class No Acknowledgement, trigger "DB302_HMI_Faults_Carrier62_Faults_0" bit 8
   3978: 'Carrier 62 Safe Output Card Fault', class No Acknowledgement, trigger "DB302_HMI_Faults_Carrier62_Faults_0" bit 9
   3979: 'Carrier 62 Standard Input Card Fault', class No Acknowledgement, trigger "DB302_HMI_Faults_Carrier62_Faults_0" bit 10
   3980: 'Carrier 62 Standard Output Card Fault', class No Acknowledgement, trigger "DB302_HMI_Faults_Carrier62_Faults_0" bit 11
   3981: 'Carrier 62 Encoder Position Fault', class No Acknowledgement, trigger "DB302_HMI_Faults_Carrier62_Faults_0" bit 12
   3982: 'Carrier 62 Encoder Internal Error', class No Acknowledgement, trigger "DB302_HMI_Faults_Carrier62_Faults_0" bit 13
   3983: 'Carrier 62 Encoder Comm Fault', class No Acknowledgement, trigger "DB302_HMI_Faults_Carrier62_Faults_0" bit 14
   3984: 'Carrier 62 HMI Comm Fault', class No Acknowledgement, trigger "DB302_HMI_Faults_Carrier62_Faults_0" bit 15
   3985: 'Carrier 62 Crash Detection Fault', class No Acknowledgement, trigger "DB302_HMI_Faults_Carrier62_Faults_1" bit 0
   3986: 'Carrier 62 Carrier Number Invalid', class No Acknowledgement, trigger "DB302_HMI_Faults_Carrier62_Faults_1" bit 1
   3987: 'Carrier 62 Drive: PROFINET configuration error', class No Acknowledgement, trigger "DB302_HMI_Faults_Carrier62_Faults_1" bit 2
   3988: 'Carrier 62 Drive: Error internal communications', class No Acknowledgement, trigger "DB302_HMI_Faults_Carrier62_Faults_1" bit 3
   3989: 'Carrier 62 Drive: Motor overtemperature', class No Acknowledgement, trigger "DB302_HMI_Faults_Carrier62_Faults_1" bit 4
   3990: 'Carrier 62 Drive: Motor overcurrent', class No Acknowledgement, trigger "DB302_HMI_Faults_Carrier62_Faults_1" bit 5
   3991: 'Carrier 62 Drive: Infeed or power unit not ready', class No Acknowledgement, trigger "DB302_HMI_Faults_Carrier62_Faults_1" bit 6
   3992: 'Carrier 62 Drive: Short-circuit/ground fault detected', class No Acknowledgement, trigger "DB302_HMI_Faults_Carrier62_Faults_1" bit 7
   3993: 'Carrier 62 Drive: PROFINET Setpoint timeout', class No Acknowledgement, trigger "DB302_HMI_Faults_Carrier62_Faults_1" bit 8
   3994: 'Carrier 62 Power unit: Overcurrent', class No Acknowledgement, trigger "DB302_HMI_Faults_Carrier62_Faults_1" bit 9
   3995: 'Carrier 62 Power unit: DC link voltage overvoltage', class No Acknowledgement, trigger "DB302_HMI_Faults_Carrier62_Faults_1" bit 10
   3996: 'Carrier 62 Power unit: DC link voltage undervoltage', class No Acknowledgement, trigger "DB302_HMI_Faults_Carrier62_Faults_1" bit 11
   3997: 'Carrier 62 Power unit: Line phase failure in main circuit', class No Acknowledgement, trigger "DB302_HMI_Faults_Carrier62_Faults_1" bit 12
   3998: 'Carrier 62 Power unit: Phase failure motor cable', class No Acknowledgement, trigger "DB302_HMI_Faults_Carrier62_Faults_1" bit 13
   3999: 'Carrier 62 Power unit: Ground fault', class No Acknowledgement, trigger "DB302_HMI_Faults_Carrier62_Faults_1" bit 14
   4000: 'Spare_Fault_4000', class No Acknowledgement, trigger "DB302_HMI_Faults_Carrier62_Faults_1" bit 15
   4001: 'Carrier 62 Motion Off Fault', class No Acknowledgement, trigger "DB302_HMI_Faults_Carrier62_Faults_2" bit 0
   4002: 'Carrier 62 Motion On Fault', class No Acknowledgement, trigger "DB302_HMI_Faults_Carrier62_Faults_2" bit 1
   4003: 'Carrier 62 Spacing Fault', class No Acknowledgement, trigger "DB302_HMI_Faults_Carrier62_Faults_2" bit 2
   4004: 'Carrier 62 Duplicate Carrier Number Fault', class No Acknowledgement, trigger "DB302_HMI_Faults_Carrier62_Faults_2" bit 3
   4005: 'Spare_Fault_4005', class No Acknowledgement, trigger "DB302_HMI_Faults_Carrier62_Faults_2" bit 4
   4006: 'Spare_Fault_4006', class No Acknowledgement, trigger "DB302_HMI_Faults_Carrier62_Faults_2" bit 5
   4007: 'Spare_Fault_4007', class No Acknowledgement, trigger "DB302_HMI_Faults_Carrier62_Faults_2" bit 6
   4008: 'Spare_Fault_4008', class No Acknowledgement, trigger "DB302_HMI_Faults_Carrier62_Faults_2" bit 7
   4009: 'Spare_Fault_4009', class No Acknowledgement, trigger "DB302_HMI_Faults_Carrier62_Faults_2" bit 8
   4010: 'Spare_Fault_4010', class No Acknowledgement, trigger "DB302_HMI_Faults_Carrier62_Faults_2" bit 9
   4011: 'Spare_Fault_4011', class No Acknowledgement, trigger "DB302_HMI_Faults_Carrier62_Faults_2" bit 10
   4012: 'Spare_Fault_4012', class No Acknowledgement, trigger "DB302_HMI_Faults_Carrier62_Faults_2" bit 11
   4013: 'Spare_Fault_4013', class No Acknowledgement, trigger "DB302_HMI_Faults_Carrier62_Faults_2" bit 12
   4014: 'Spare_Fault_4014', class No Acknowledgement, trigger "DB302_HMI_Faults_Carrier62_Faults_2" bit 13
   4015: 'Spare_Fault_4015', class No Acknowledgement, trigger "DB302_HMI_Faults_Carrier62_Faults_2" bit 14
   4016: 'Spare_Fault_4016', class No Acknowledgement, trigger "DB302_HMI_Faults_Carrier62_Faults_2" bit 15
   4017: 'Spare_Fault_4017', class No Acknowledgement, trigger "DB302_HMI_Faults_Carrier62_Faults_3" bit 0
   4018: 'Spare_Fault_4018', class No Acknowledgement, trigger "DB302_HMI_Faults_Carrier62_Faults_3" bit 1
   4019: 'Spare_Fault_4019', class No Acknowledgement, trigger "DB302_HMI_Faults_Carrier62_Faults_3" bit 2
   4020: 'Spare_Fault_4020', class No Acknowledgement, trigger "DB302_HMI_Faults_Carrier62_Faults_3" bit 3
   4021: 'Spare_Fault_4021', class No Acknowledgement, trigger "DB302_HMI_Faults_Carrier62_Faults_3" bit 4
   4022: 'Spare_Fault_4022', class No Acknowledgement, trigger "DB302_HMI_Faults_Carrier62_Faults_3" bit 5
   4023: 'Spare_Fault_4023', class No Acknowledgement, trigger "DB302_HMI_Faults_Carrier62_Faults_3" bit 6
   4024: 'Spare_Fault_4024', class No Acknowledgement, trigger "DB302_HMI_Faults_Carrier62_Faults_3" bit 7
   4025: 'Spare_Fault_4025', class No Acknowledgement, trigger "DB302_HMI_Faults_Carrier62_Faults_3" bit 8
   4026: 'Spare_Fault_4026', class No Acknowledgement, trigger "DB302_HMI_Faults_Carrier62_Faults_3" bit 9
   4027: 'Spare_Fault_4027', class No Acknowledgement, trigger "DB302_HMI_Faults_Carrier62_Faults_3" bit 10
   4028: 'Spare_Fault_4028', class No Acknowledgement, trigger "DB302_HMI_Faults_Carrier62_Faults_3" bit 11
   4029: 'Spare_Fault_4029', class No Acknowledgement, trigger "DB302_HMI_Faults_Carrier62_Faults_3" bit 12
   4030: 'Spare_Fault_4030', class No Acknowledgement, trigger "DB302_HMI_Faults_Carrier62_Faults_3" bit 13
   4031: 'Spare_Fault_4031', class No Acknowledgement, trigger "DB302_HMI_Faults_Carrier62_Faults_3" bit 14
   4032: 'Spare_Fault_4032', class No Acknowledgement, trigger "DB302_HMI_Faults_Carrier62_Faults_3" bit 15
   4033: 'Carrier 63 Disconnect Open Power Fault DI11.0', class No Acknowledgement, trigger "DB302_HMI_Faults_Carrier63_Faults_0" bit 0
   4034: 'Carrier 63 Drive Profinet Comm Fault', class No Acknowledgement, trigger "DB302_HMI_Faults_Carrier63_Faults_0" bit 1
   4035: 'Carrier 63 Production Stop Not Reset', class No Acknowledgement, trigger "DB302_HMI_Faults_Carrier63_Faults_0" bit 2
   4036: 'Carrier 63 CB02122 Tripped', class No Acknowledgement, trigger "DB302_HMI_Faults_Carrier63_Faults_0" bit 3
   4037: 'Carrier 63 CB02123 Tripped', class No Acknowledgement, trigger "DB302_HMI_Faults_Carrier63_Faults_0" bit 4
   4038: 'Carrier 63 AUX1 CB Tripped', class No Acknowledgement, trigger "DB302_HMI_Faults_Carrier63_Faults_0" bit 5
   4039: 'Carrier 63 AUX2 CB Tripped', class No Acknowledgement, trigger "DB302_HMI_Faults_Carrier63_Faults_0" bit 6
   4040: 'Carrier 63 PLC Not Communicating', class No Acknowledgement, trigger "DB302_HMI_Faults_Carrier63_Faults_0" bit 7
   4041: 'Carrier 63 Safe Input Card Fault', class No Acknowledgement, trigger "DB302_HMI_Faults_Carrier63_Faults_0" bit 8
   4042: 'Carrier 63 Safe Output Card Fault', class No Acknowledgement, trigger "DB302_HMI_Faults_Carrier63_Faults_0" bit 9
   4043: 'Carrier 63 Standard Input Card Fault', class No Acknowledgement, trigger "DB302_HMI_Faults_Carrier63_Faults_0" bit 10
   4044: 'Carrier 63 Standard Output Card Fault', class No Acknowledgement, trigger "DB302_HMI_Faults_Carrier63_Faults_0" bit 11
   4045: 'Carrier 63 Encoder Position Fault', class No Acknowledgement, trigger "DB302_HMI_Faults_Carrier63_Faults_0" bit 12
   4046: 'Carrier 63 Encoder Internal Error', class No Acknowledgement, trigger "DB302_HMI_Faults_Carrier63_Faults_0" bit 13
   4047: 'Carrier 63 Encoder Comm Fault', class No Acknowledgement, trigger "DB302_HMI_Faults_Carrier63_Faults_0" bit 14
   4048: 'Carrier 63 HMI Comm Fault', class No Acknowledgement, trigger "DB302_HMI_Faults_Carrier63_Faults_0" bit 15
   4049: 'Carrier 63 Crash Detection Fault', class No Acknowledgement, trigger "DB302_HMI_Faults_Carrier63_Faults_1" bit 0
   4050: 'Carrier 63 Carrier Number Invalid', class No Acknowledgement, trigger "DB302_HMI_Faults_Carrier63_Faults_1" bit 1
   4051: 'Carrier 63 Drive: PROFINET configuration error', class No Acknowledgement, trigger "DB302_HMI_Faults_Carrier63_Faults_1" bit 2
   4052: 'Carrier 63 Drive: Error internal communications', class No Acknowledgement, trigger "DB302_HMI_Faults_Carrier63_Faults_1" bit 3
   4053: 'Carrier 63 Drive: Motor overtemperature', class No Acknowledgement, trigger "DB302_HMI_Faults_Carrier63_Faults_1" bit 4
   4054: 'Carrier 63 Drive: Motor overcurrent', class No Acknowledgement, trigger "DB302_HMI_Faults_Carrier63_Faults_1" bit 5
   4055: 'Carrier 63 Drive: Infeed or power unit not ready', class No Acknowledgement, trigger "DB302_HMI_Faults_Carrier63_Faults_1" bit 6
   4056: 'Carrier 63 Drive: Short-circuit/ground fault detected', class No Acknowledgement, trigger "DB302_HMI_Faults_Carrier63_Faults_1" bit 7
   4057: 'Carrier 63 Drive: PROFINET Setpoint timeout', class No Acknowledgement, trigger "DB302_HMI_Faults_Carrier63_Faults_1" bit 8
   4058: 'Carrier 63 Power unit: Overcurrent', class No Acknowledgement, trigger "DB302_HMI_Faults_Carrier63_Faults_1" bit 9
   4059: 'Carrier 63 Power unit: DC link voltage overvoltage', class No Acknowledgement, trigger "DB302_HMI_Faults_Carrier63_Faults_1" bit 10
   4060: 'Carrier 63 Power unit: DC link voltage undervoltage', class No Acknowledgement, trigger "DB302_HMI_Faults_Carrier63_Faults_1" bit 11
   4061: 'Carrier 63 Power unit: Line phase failure in main circuit', class No Acknowledgement, trigger "DB302_HMI_Faults_Carrier63_Faults_1" bit 12
   4062: 'Carrier 63 Power unit: Phase failure motor cable', class No Acknowledgement, trigger "DB302_HMI_Faults_Carrier63_Faults_1" bit 13
   4063: 'Carrier 63 Power unit: Ground fault', class No Acknowledgement, trigger "DB302_HMI_Faults_Carrier63_Faults_1" bit 14
   4064: 'Spare_Fault_4064', class No Acknowledgement, trigger "DB302_HMI_Faults_Carrier63_Faults_1" bit 15
   4065: 'Carrier 63 Motion Off Fault', class No Acknowledgement, trigger "DB302_HMI_Faults_Carrier63_Faults_2" bit 0
   4066: 'Carrier 63 Motion On Fault', class No Acknowledgement, trigger "DB302_HMI_Faults_Carrier63_Faults_2" bit 1
